REGION Network 9
   RUNG wire#powerrail
      Move(in := #AccumZnSpacing, out1 => #AccumSpacingEcho)
      Move(in := #ProductZoneSpacing, out1 => #ProdZoneSpacingEcho)
   END_RUNG
   // the same network as SCL:
   #AccumSpacingEcho := #AccumZnSpacing;
   #ProdZoneSpacingEcho := #ProductZoneSpacing;
END_REGION

REGION Network 10
   RUNG wire#powerrail
      { S7_Templates := "SrcType := Int" } NE_Contact(in1 := "EMS".Zone[#Zone].CarrierZnStatus[#MaxCarriers].CarrierNumber, in2 := 0)
      Coil( #ZoneFull )
   END_RUNG
   // the same network as SCL:
   #ZoneFull := "EMS".Zone[#Zone].CarrierZnStatus[#MaxCarriers].CarrierNumber <> 0;
END_REGION

REGION Network 11
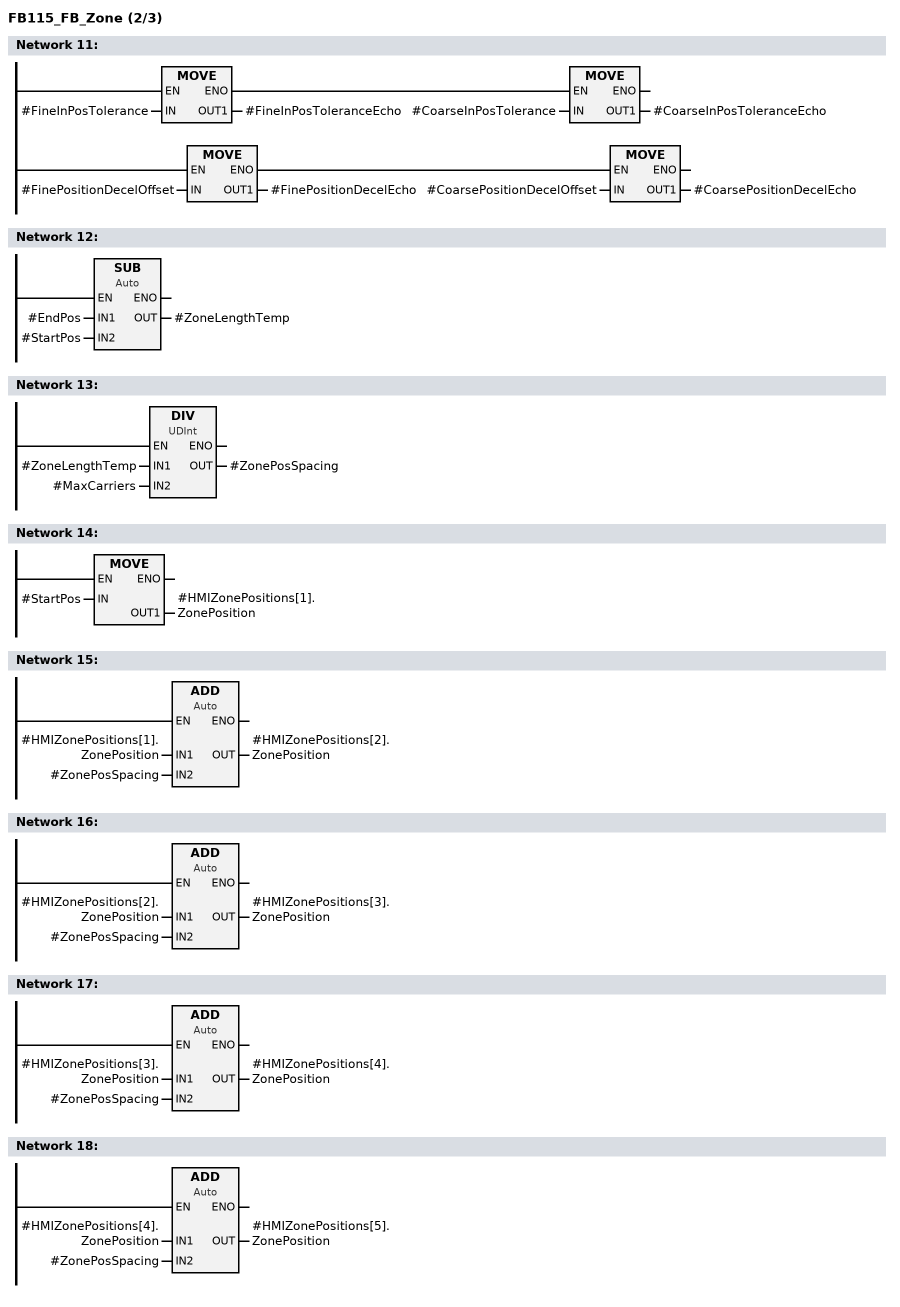
   RUNG wire#powerrail
      Move(in := #FineInPosTolerance, out1 => #FineInPosToleranceEcho)
      Move(in := #CoarseInPosTolerance, out1 => #CoarseInPosToleranceEcho)
   END_RUNG
   RUNG wire#powerrail
      Move(in := #FinePositionDecelOffset, out1 => #FinePositionDecelEcho)
      Move(in := #CoarsePositionDecelOffset, out1 => #CoarsePositionDecelEcho)
   END_RUNG
   // the same network as SCL:
   #FineInPosToleranceEcho := #FineInPosTolerance;
   #CoarseInPosToleranceEcho := #CoarseInPosTolerance;
   #FinePositionDecelEcho := #FinePositionDecelOffset;
   #CoarsePositionDecelEcho := #CoarsePositionDecelOffset;
END_REGION

REGION Network 12
   RUNG wire#powerrail
      Sub(in1 := #EndPos, in2 := #StartPos, out => #ZoneLengthTemp)
   END_RUNG
   // the same network as SCL:
   #ZoneLengthTemp := #EndPos - #StartPos;
END_REGION

REGION Network 13
   RUNG wire#powerrail
      { S7_Templates := "SrcType := UDInt" } Div(in1 := #ZoneLengthTemp, in2 := #MaxCarriers, out => #ZonePosSpacing)
   END_RUNG
   // the same network as SCL:
   #ZonePosSpacing := #ZoneLengthTemp / #MaxCarriers;
END_REGION

REGION Network 14
   RUNG wire#powerrail
      Move(in := #StartPos, out1 => #HMIZonePositions[1].ZonePosition)
   END_RUNG
   // the same network as SCL:
   #HMIZonePositions[1].ZonePosition := #StartPos;
END_REGION

REGION Network 15
   RUNG wire#powerrail
      Add(in1 := #HMIZonePositions[1].ZonePosition, in2 := #ZonePosSpacing, out => #HMIZonePositions[2].ZonePosition)
   END_RUNG
   // the same network as SCL:
   #HMIZonePositions[2].ZonePosition := #HMIZonePositions[1].ZonePosition + #ZonePosSpacing;
END_REGION

REGION Network 16
   RUNG wire#powerrail
      Add(in1 := #HMIZonePositions[2].ZonePosition, in2 := #ZonePosSpacing, out => #HMIZonePositions[3].ZonePosition)
   END_RUNG
   // the same network as SCL:
   #HMIZonePositions[3].ZonePosition := #HMIZonePositions[2].ZonePosition + #ZonePosSpacing;
END_REGION

REGION Network 17
   RUNG wire#powerrail
      Add(in1 := #HMIZonePositions[3].ZonePosition, in2 := #ZonePosSpacing, out => #HMIZonePositions[4].ZonePosition)
   END_RUNG
   // the same network as SCL:
   #HMIZonePositions[4].ZonePosition := #HMIZonePositions[3].ZonePosition + #ZonePosSpacing;
END_REGION

REGION Network 18
   RUNG wire#powerrail
      Add(in1 := #HMIZonePositions[4].ZonePosition, in2 := #ZonePosSpacing, out => #HMIZonePositions[5].ZonePosition)
   END_RUNG
   // the same network as SCL:
   #HMIZonePositions[5].ZonePosition := #HMIZonePositions[4].ZonePosition + #ZonePosSpacing;
END_REGION

REGION Network 19
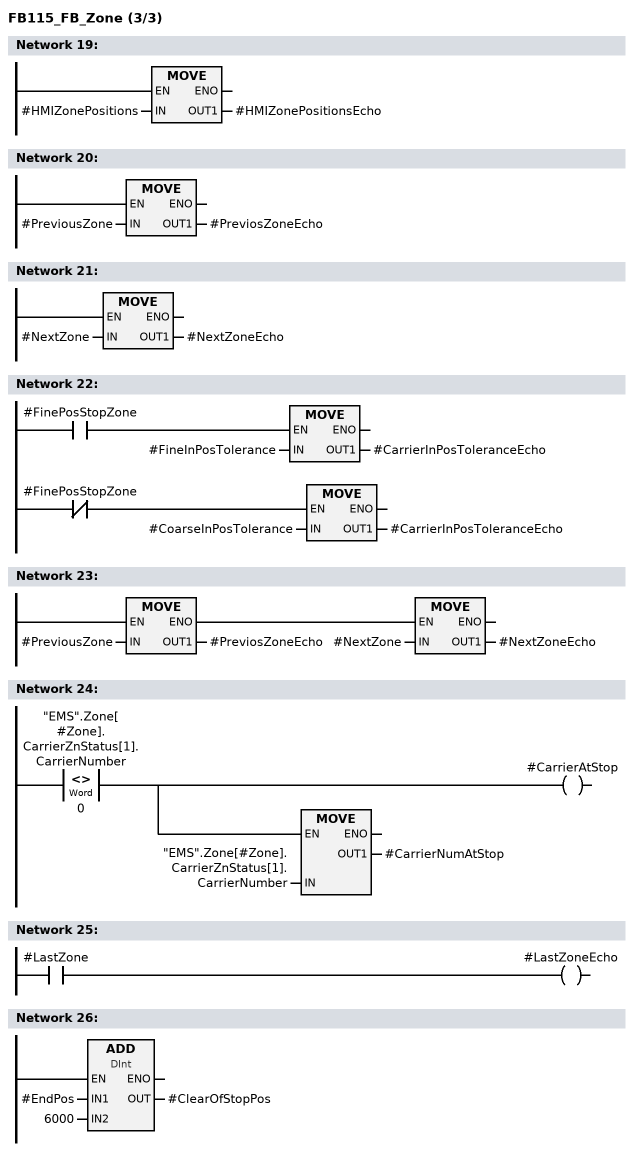
   RUNG wire#powerrail
      Move(in := #HMIZonePositions, out1 => #HMIZonePositionsEcho)
   END_RUNG
   // the same network as SCL:
   #HMIZonePositionsEcho := #HMIZonePositions;
END_REGION

REGION Network 20
   RUNG wire#powerrail
      Move(in := #PreviousZone, out1 => #PreviosZoneEcho)
   END_RUNG
   // the same network as SCL:
   #PreviosZoneEcho := #PreviousZone;
END_REGION

REGION Network 21
   RUNG wire#powerrail
      Move(in := #NextZone, out1 => #NextZoneEcho)
   END_RUNG
   // the same network as SCL:
   #NextZoneEcho := #NextZone;
END_REGION

REGION Network 22
   RUNG wire#powerrail
      Contact( #FinePosStopZone )
      Move(in := #FineInPosTolerance, out1 => #CarrierInPosToleranceEcho)
   END_RUNG
   RUNG wire#powerrail
      I_Contact( #FinePosStopZone )
      Move(in := #CoarseInPosTolerance, out1 => #CarrierInPosToleranceEcho)
   END_RUNG
   // the same network as SCL:
   IF #FinePosStopZone THEN #CarrierInPosToleranceEcho := #FineInPosTolerance; END_IF;
   IF NOT #FinePosStopZone THEN #CarrierInPosToleranceEcho := #CoarseInPosTolerance; END_IF;
END_REGION

REGION Network 23
   RUNG wire#powerrail
      Move(in := #PreviousZone, out1 => #PreviosZoneEcho)
      Move(in := #NextZone, out1 => #NextZoneEcho)
   END_RUNG
   // the same network as SCL:
   #PreviosZoneEcho := #PreviousZone;
   #NextZoneEcho := #NextZone;
END_REGION

REGION Network 24
   RUNG wire#powerrail
      { S7_Templates := "SrcType := Word" } NE_Contact(in1 := "EMS".Zone[#Zone].CarrierZnStatus[1].CarrierNumber, in2 := 0)
      wire#w1
      Coil( #CarrierAtStop )
   END_RUNG
   RUNG wire#w1
      Move(in := "EMS".Zone[#Zone].CarrierZnStatus[1].CarrierNumber, out1 => #CarrierNumAtStop)
   END_RUNG
   // the same network as SCL:
   #CarrierAtStop := "EMS".Zone[#Zone].CarrierZnStatus[1].CarrierNumber <> 0;
   IF #CarrierAtStop THEN #CarrierNumAtStop := "EMS".Zone[#Zone].CarrierZnStatus[1].CarrierNumber; END_IF;
END_REGION

REGION Network 25
   RUNG wire#powerrail
      Contact( #LastZone )
      Coil( #LastZoneEcho )
   END_RUNG
   // the same network as SCL:
   #LastZoneEcho := #LastZone;
END_REGION

REGION Network 26
   RUNG wire#powerrail
      { S7_Templates := "SrcType := DInt" } Add(in1 := #EndPos, in2 := 6000, out => #ClearOfStopPos)
   END_RUNG
   // the same network as SCL:
   #ClearOfStopPos := #EndPos + 6000;
END_REGION
END_FUNCTION_BLOCK

FUNCTION_BLOCK "FB116_FB_ZonePositionArrayTrafficCop"   // FB116, LAD
{ S7_Optimized_Access := 'FALSE' }
VERSION : 0.1
   VAR_INPUT
      Zone : Int := 1;
      CarrierZnArrayPos : Int;
   END_VAR
   VAR_OUTPUT
      MoveFwd : Bool;
      Speed : Word;
      TCZnPosnArray : "UDT_TrafficCopZoneStructure";
   END_VAR
   VAR
      CarNumZnPos : Array[0..99] of Int;
      TrafficCopCarrierZnBufferOut : Array[0..30] of "UDT_TrafficCop";
      "Zn-Pos2CarrierNumTemp" : Int;
      Zone1TrafficCopStructure : Struct
         CommandPosition : Word;
         InPositionTolerance : Word;
         CommandPositionUpperLimit : Word;
         CommandPositionLowerLimit : Word;
         AtCommandPos : Bool;
      END_STRUCT;
      SectionComment : Bool;
      NextCarrierZnArrayPos : Int;
   END_VAR
BEGIN

REGION Network 1: Section Comment-Section Logic for Current Carrier number in Position 1 thru Max Carrier in Zone Position Array
   // Section Logic for Current Carrier number in Position 1 - Max Carrier in Zone Position Array
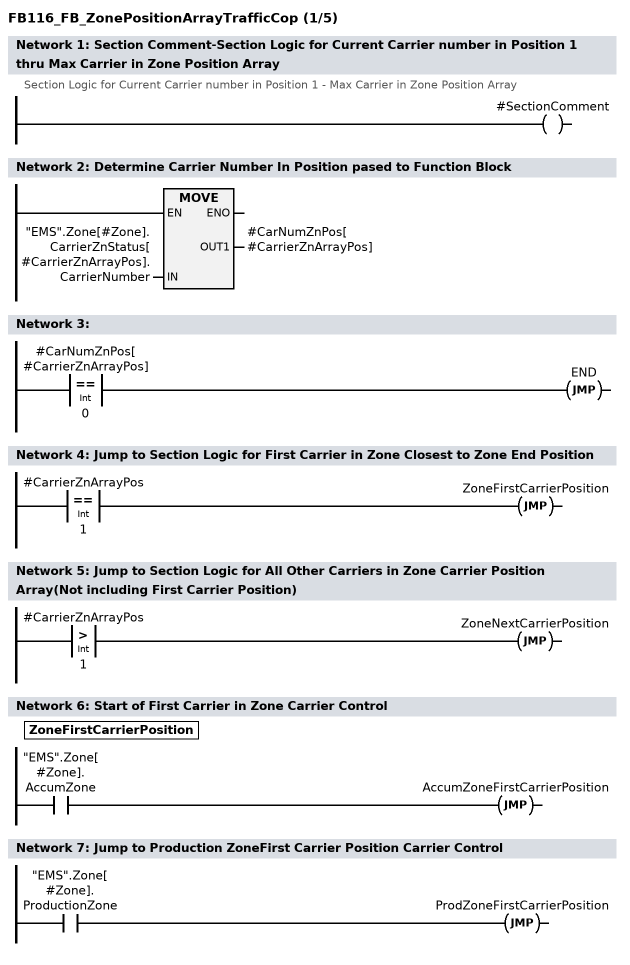
   RUNG wire#powerrail
      Coil( #SectionComment )
   END_RUNG
   // the same network as SCL:
   #SectionComment := TRUE;
END_REGION

REGION Network 2: Determine Carrier Number In Position pased to Function Block
   RUNG wire#powerrail
      Move(in := "EMS".Zone[#Zone].CarrierZnStatus[#CarrierZnArrayPos].CarrierNumber, out1 => #CarNumZnPos[#CarrierZnArrayPos])
   END_RUNG
   // the same network as SCL:
   #CarNumZnPos[#CarrierZnArrayPos] := "EMS".Zone[#Zone].CarrierZnStatus[#CarrierZnArrayPos].CarrierNumber;
END_REGION

REGION Network 3
   RUNG wire#powerrail
      { S7_Templates := "SrcType := Int" } EQ_Contact(in1 := #CarNumZnPos[#CarrierZnArrayPos], in2 := 0)
      JumpCoil( END )
   END_RUNG
   // the same network as SCL:
   IF #CarNumZnPos[#CarrierZnArrayPos] = 0 THEN GOTO END; END_IF;
END_REGION

REGION Network 4: Jump to Section Logic for First Carrier in Zone Closest to Zone End Position
   RUNG wire#powerrail
      { S7_Templates := "SrcType := Int" } EQ_Contact(in1 := #CarrierZnArrayPos, in2 := 1)
      JumpCoil( ZoneFirstCarrierPosition )
   END_RUNG
   // the same network as SCL:
   IF #CarrierZnArrayPos = 1 THEN GOTO ZoneFirstCarrierPosition; END_IF;
END_REGION

REGION Network 5: Jump to Section Logic for All Other Carriers in Zone Carrier Position Array(Not including First Carrier Position)
   RUNG wire#powerrail
      { S7_Templates := "SrcType := Int" } GT_Contact(in1 := #CarrierZnArrayPos, in2 := 1)
      JumpCoil( ZoneNextCarrierPosition )
   END_RUNG
   // the same network as SCL:
   IF #CarrierZnArrayPos > 1 THEN GOTO ZoneNextCarrierPosition; END_IF;
END_REGION

REGION Network 6: Start of First Carrier in Zone Carrier Control
   Label( ZoneFirstCarrierPosition )
   RUNG wire#powerrail
      Contact( "EMS".Zone[#Zone].AccumZone )
      JumpCoil( AccumZoneFirstCarrierPosition )
   END_RUNG
   // the same network as SCL:
   ZoneFirstCarrierPosition:
   IF "EMS".Zone[#Zone].AccumZone THEN GOTO AccumZoneFirstCarrierPosition; END_IF;
END_REGION

REGION Network 7: Jump to Production ZoneFirst Carrier Position Carrier Control
   RUNG wire#powerrail
      Contact( "EMS".Zone[#Zone].ProductionZone )
      JumpCoil( ProdZoneFirstCarrierPosition )
   END_RUNG
   // the same network as SCL:
   IF "EMS".Zone[#Zone].ProductionZone THEN GOTO ProdZoneFirstCarrierPosition; END_IF;
END_REGION

REGION Network 8: Position Carrier Control First Carrier in Accumulation Zone
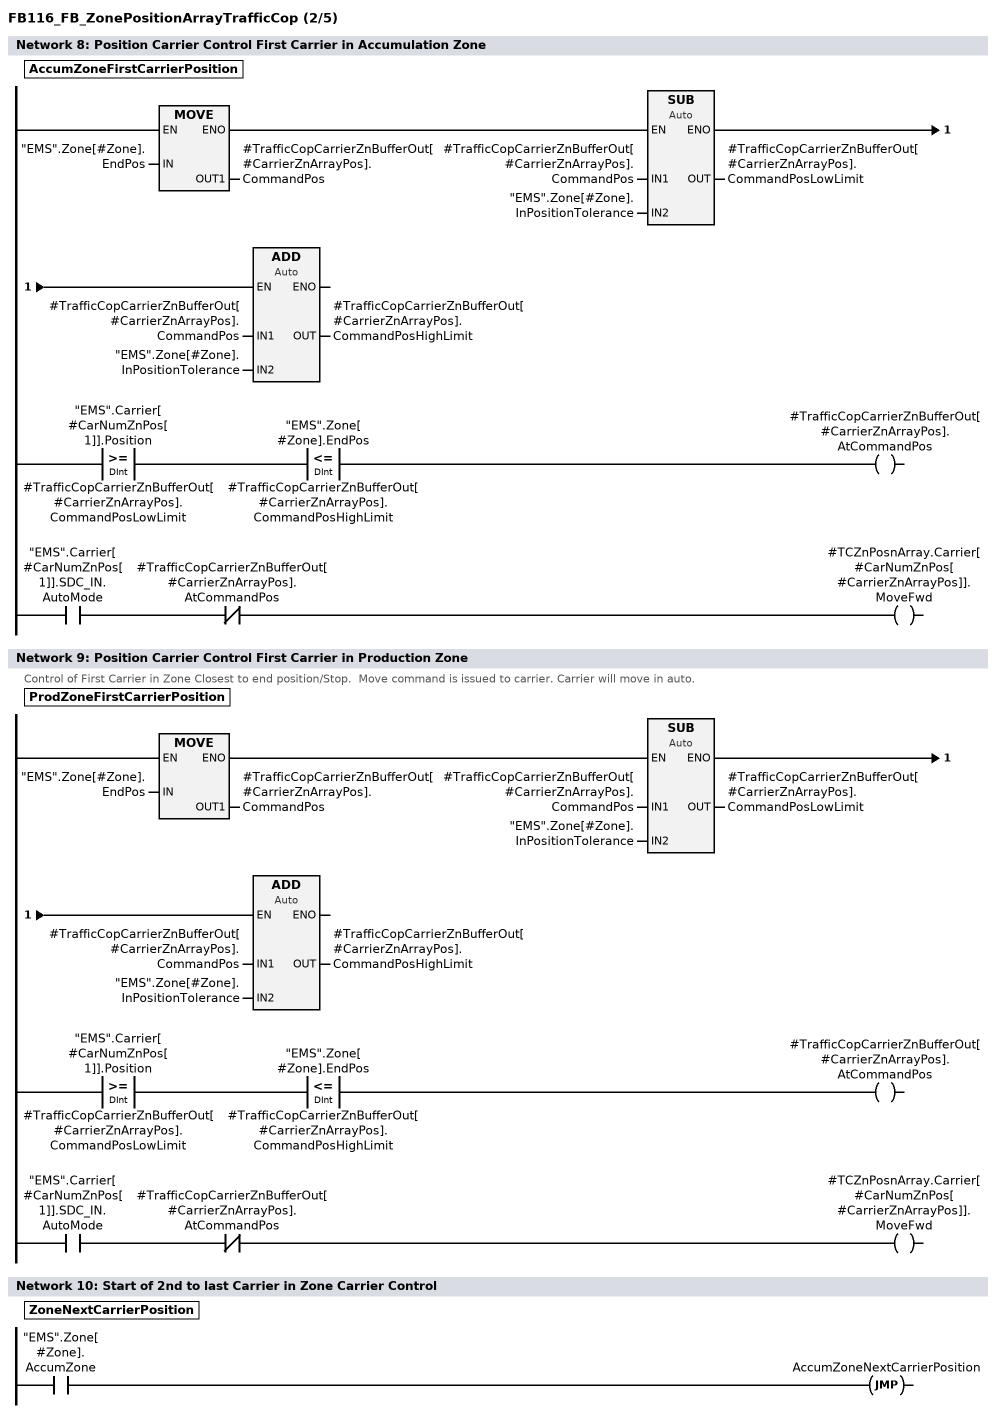
   Label( AccumZoneFirstCarrierPosition )
   RUNG wire#powerrail
      Move(in := "EMS".Zone[#Zone].EndPos, out1 => #TrafficCopCarrierZnBufferOut[#CarrierZnArrayPos].CommandPos)
      Sub(in1 := #TrafficCopCarrierZnBufferOut[#CarrierZnArrayPos].CommandPos, in2 := "EMS".Zone[#Zone].InPositionTolerance, out => #TrafficCopCarrierZnBufferOut[#CarrierZnArrayPos].CommandPosLowLimit)
      Add(in1 := #TrafficCopCarrierZnBufferOut[#CarrierZnArrayPos].CommandPos, in2 := "EMS".Zone[#Zone].InPositionTolerance, out => #TrafficCopCarrierZnBufferOut[#CarrierZnArrayPos].CommandPosHighLimit)
   END_RUNG
   RUNG wire#powerrail
      { S7_Templates := "SrcType := DInt" } GE_Contact(in1 := "EMS".Carrier[#CarNumZnPos[1]].Position, in2 := #TrafficCopCarrierZnBufferOut[#CarrierZnArrayPos].CommandPosLowLimit)
      { S7_Templates := "SrcType := DInt" } LE_Contact(in1 := "EMS".Zone[#Zone].EndPos, in2 := #TrafficCopCarrierZnBufferOut[#CarrierZnArrayPos].CommandPosHighLimit)
      Coil( #TrafficCopCarrierZnBufferOut[#CarrierZnArrayPos].AtCommandPos )
   END_RUNG
   RUNG wire#powerrail
      Contact( "EMS".Carrier[#CarNumZnPos[1]].SDC_IN.AutoMode )
      I_Contact( #TrafficCopCarrierZnBufferOut[#CarrierZnArrayPos].AtCommandPos )
      Coil( #TCZnPosnArray.Carrier[#CarNumZnPos[#CarrierZnArrayPos]].MoveFwd )
   END_RUNG
   // the same network as SCL:
   AccumZoneFirstCarrierPosition:
   #TrafficCopCarrierZnBufferOut[#CarrierZnArrayPos].CommandPos := "EMS".Zone[#Zone].EndPos;
   #TrafficCopCarrierZnBufferOut[#CarrierZnArrayPos].CommandPosLowLimit := #TrafficCopCarrierZnBufferOut[#CarrierZnArrayPos].CommandPos - "EMS".Zone[#Zone].InPositionTolerance;
   #TrafficCopCarrierZnBufferOut[#CarrierZnArrayPos].CommandPosHighLimit := #TrafficCopCarrierZnBufferOut[#CarrierZnArrayPos].CommandPos + "EMS".Zone[#Zone].InPositionTolerance;
   #TrafficCopCarrierZnBufferOut[#CarrierZnArrayPos].AtCommandPos := ("EMS".Carrier[#CarNumZnPos[1]].Position >= #TrafficCopCarrierZnBufferOut[#CarrierZnArrayPos].CommandPosLowLimit) AND ("EMS".Zone[#Zone].EndPos <= #TrafficCopCarrierZnBufferOut[#CarrierZnArrayPos].CommandPosHighLimit);
   #TCZnPosnArray.Carrier[#CarNumZnPos[#CarrierZnArrayPos]].MoveFwd := "EMS".Carrier[#CarNumZnPos[1]].SDC_IN.AutoMode AND NOT #TrafficCopCarrierZnBufferOut[#CarrierZnArrayPos].AtCommandPos;
END_REGION

REGION Network 9: Position Carrier Control First Carrier in Production Zone
   // Control of First Carrier in Zone Closest to end position/Stop.  Move command is issued to carrier. Carrier will move in auto.
   Label( ProdZoneFirstCarrierPosition )
   RUNG wire#powerrail
      Move(in := "EMS".Zone[#Zone].EndPos, out1 => #TrafficCopCarrierZnBufferOut[#CarrierZnArrayPos].CommandPos)
      Sub(in1 := #TrafficCopCarrierZnBufferOut[#CarrierZnArrayPos].CommandPos, in2 := "EMS".Zone[#Zone].InPositionTolerance, out => #TrafficCopCarrierZnBufferOut[#CarrierZnArrayPos].CommandPosLowLimit)
      Add(in1 := #TrafficCopCarrierZnBufferOut[#CarrierZnArrayPos].CommandPos, in2 := "EMS".Zone[#Zone].InPositionTolerance, out => #TrafficCopCarrierZnBufferOut[#CarrierZnArrayPos].CommandPosHighLimit)
   END_RUNG
   RUNG wire#powerrail
      { S7_Templates := "SrcType := DInt" } GE_Contact(in1 := "EMS".Carrier[#CarNumZnPos[1]].Position, in2 := #TrafficCopCarrierZnBufferOut[#CarrierZnArrayPos].CommandPosLowLimit)
      { S7_Templates := "SrcType := DInt" } LE_Contact(in1 := "EMS".Zone[#Zone].EndPos, in2 := #TrafficCopCarrierZnBufferOut[#CarrierZnArrayPos].CommandPosHighLimit)
      Coil( #TrafficCopCarrierZnBufferOut[#CarrierZnArrayPos].AtCommandPos )
   END_RUNG
   RUNG wire#powerrail
      Contact( "EMS".Carrier[#CarNumZnPos[1]].SDC_IN.AutoMode )
      I_Contact( #TrafficCopCarrierZnBufferOut[#CarrierZnArrayPos].AtCommandPos )
      Coil( #TCZnPosnArray.Carrier[#CarNumZnPos[#CarrierZnArrayPos]].MoveFwd )
   END_RUNG
   // the same network as SCL:
   ProdZoneFirstCarrierPosition:
   #TrafficCopCarrierZnBufferOut[#CarrierZnArrayPos].CommandPos := "EMS".Zone[#Zone].EndPos;
   #TrafficCopCarrierZnBufferOut[#CarrierZnArrayPos].CommandPosLowLimit := #TrafficCopCarrierZnBufferOut[#CarrierZnArrayPos].CommandPos - "EMS".Zone[#Zone].InPositionTolerance;
   #TrafficCopCarrierZnBufferOut[#CarrierZnArrayPos].CommandPosHighLimit := #TrafficCopCarrierZnBufferOut[#CarrierZnArrayPos].CommandPos + "EMS".Zone[#Zone].InPositionTolerance;
   #TrafficCopCarrierZnBufferOut[#CarrierZnArrayPos].AtCommandPos := ("EMS".Carrier[#CarNumZnPos[1]].Position >= #TrafficCopCarrierZnBufferOut[#CarrierZnArrayPos].CommandPosLowLimit) AND ("EMS".Zone[#Zone].EndPos <= #TrafficCopCarrierZnBufferOut[#CarrierZnArrayPos].CommandPosHighLimit);
   #TCZnPosnArray.Carrier[#CarNumZnPos[#CarrierZnArrayPos]].MoveFwd := "EMS".Carrier[#CarNumZnPos[1]].SDC_IN.AutoMode AND NOT #TrafficCopCarrierZnBufferOut[#CarrierZnArrayPos].AtCommandPos;
END_REGION

REGION Network 10: Start of 2nd to last Carrier in Zone Carrier Control
   Label( ZoneNextCarrierPosition )
   RUNG wire#powerrail
      Contact( "EMS".Zone[#Zone].AccumZone )
      JumpCoil( AccumZoneNextCarrierPosition )
   END_RUNG
   // the same network as SCL:
   ZoneNextCarrierPosition:
   IF "EMS".Zone[#Zone].AccumZone THEN GOTO AccumZoneNextCarrierPosition; END_IF;
END_REGION

REGION Network 11: Jump to Production Zone 2nd to Last Carrier Position Carrier Control
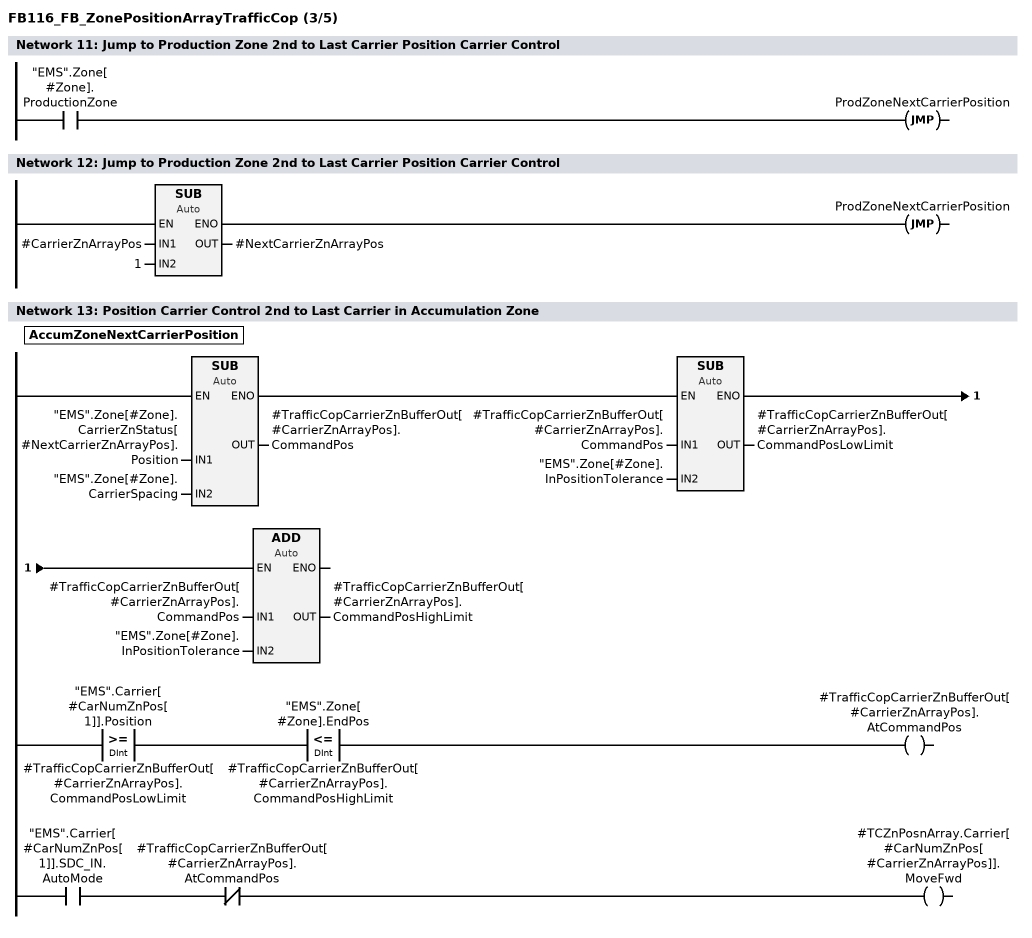
   RUNG wire#powerrail
      Contact( "EMS".Zone[#Zone].ProductionZone )
      JumpCoil( ProdZoneNextCarrierPosition )
   END_RUNG
   // the same network as SCL:
   IF "EMS".Zone[#Zone].ProductionZone THEN GOTO ProdZoneNextCarrierPosition; END_IF;
END_REGION

REGION Network 12: Jump to Production Zone 2nd to Last Carrier Position Carrier Control
   RUNG wire#powerrail
      Sub(in1 := #CarrierZnArrayPos, in2 := 1, out => #NextCarrierZnArrayPos)
      JumpCoil( ProdZoneNextCarrierPosition )
   END_RUNG
   // the same network as SCL:
   #NextCarrierZnArrayPos := #CarrierZnArrayPos - 1;
   GOTO ProdZoneNextCarrierPosition;
END_REGION

REGION Network 13: Position Carrier Control 2nd to Last Carrier in Accumulation Zone
   Label( AccumZoneNextCarrierPosition )
   RUNG wire#powerrail
      Sub(in1 := "EMS".Zone[#Zone].CarrierZnStatus[#NextCarrierZnArrayPos].Position, in2 := "EMS".Zone[#Zone].CarrierSpacing, out => #TrafficCopCarrierZnBufferOut[#CarrierZnArrayPos].CommandPos)
      Sub(in1 := #TrafficCopCarrierZnBufferOut[#CarrierZnArrayPos].CommandPos, in2 := "EMS".Zone[#Zone].InPositionTolerance, out => #TrafficCopCarrierZnBufferOut[#CarrierZnArrayPos].CommandPosLowLimit)
      Add(in1 := #TrafficCopCarrierZnBufferOut[#CarrierZnArrayPos].CommandPos, in2 := "EMS".Zone[#Zone].InPositionTolerance, out => #TrafficCopCarrierZnBufferOut[#CarrierZnArrayPos].CommandPosHighLimit)
   END_RUNG
   RUNG wire#powerrail
      { S7_Templates := "SrcType := DInt" } GE_Contact(in1 := "EMS".Carrier[#CarNumZnPos[1]].Position, in2 := #TrafficCopCarrierZnBufferOut[#CarrierZnArrayPos].CommandPosLowLimit)
      { S7_Templates := "SrcType := DInt" } LE_Contact(in1 := "EMS".Zone[#Zone].EndPos, in2 := #TrafficCopCarrierZnBufferOut[#CarrierZnArrayPos].CommandPosHighLimit)
      Coil( #TrafficCopCarrierZnBufferOut[#CarrierZnArrayPos].AtCommandPos )
   END_RUNG
   RUNG wire#powerrail
      Contact( "EMS".Carrier[#CarNumZnPos[1]].SDC_IN.AutoMode )
      I_Contact( #TrafficCopCarrierZnBufferOut[#CarrierZnArrayPos].AtCommandPos )
      Coil( #TCZnPosnArray.Carrier[#CarNumZnPos[#CarrierZnArrayPos]].MoveFwd )
   END_RUNG
   // the same network as SCL:
   AccumZoneNextCarrierPosition:
   #TrafficCopCarrierZnBufferOut[#CarrierZnArrayPos].CommandPos := "EMS".Zone[#Zone].CarrierZnStatus[#NextCarrierZnArrayPos].Position - "EMS".Zone[#Zone].CarrierSpacing;
   #TrafficCopCarrierZnBufferOut[#CarrierZnArrayPos].CommandPosLowLimit := #TrafficCopCarrierZnBufferOut[#CarrierZnArrayPos].CommandPos - "EMS".Zone[#Zone].InPositionTolerance;
   #TrafficCopCarrierZnBufferOut[#CarrierZnArrayPos].CommandPosHighLimit := #TrafficCopCarrierZnBufferOut[#CarrierZnArrayPos].CommandPos + "EMS".Zone[#Zone].InPositionTolerance;
   #TrafficCopCarrierZnBufferOut[#CarrierZnArrayPos].AtCommandPos := ("EMS".Carrier[#CarNumZnPos[1]].Position >= #TrafficCopCarrierZnBufferOut[#CarrierZnArrayPos].CommandPosLowLimit) AND ("EMS".Zone[#Zone].EndPos <= #TrafficCopCarrierZnBufferOut[#CarrierZnArrayPos].CommandPosHighLimit);
   #TCZnPosnArray.Carrier[#CarNumZnPos[#CarrierZnArrayPos]].MoveFwd := "EMS".Carrier[#CarNumZnPos[1]].SDC_IN.AutoMode AND NOT #TrafficCopCarrierZnBufferOut[#CarrierZnArrayPos].AtCommandPos;
END_REGION

REGION Network 14: Position Carrier Control 2nd to Last Carrier in Production Zone
   // Control of 2nd to Last Carrier in Zone Move to next zone with carrier spacing
   // .  Move command is issued to carrier. Carrier will move in auto.
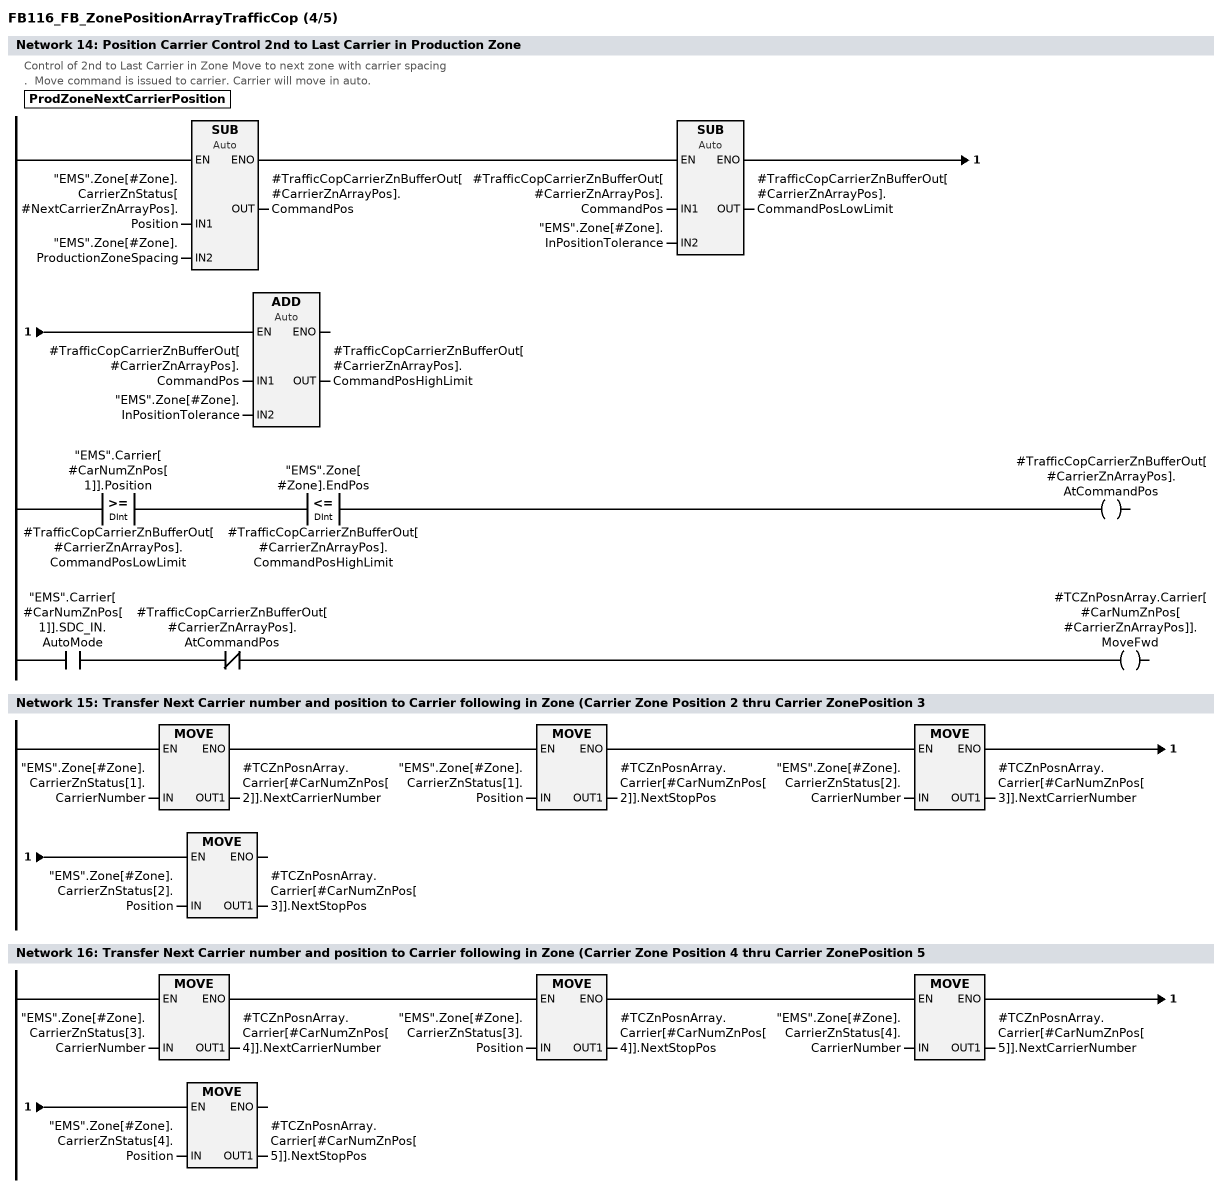
   Label( ProdZoneNextCarrierPosition )
   RUNG wire#powerrail
      Sub(in1 := "EMS".Zone[#Zone].CarrierZnStatus[#NextCarrierZnArrayPos].Position, in2 := "EMS".Zone[#Zone].ProductionZoneSpacing, out => #TrafficCopCarrierZnBufferOut[#CarrierZnArrayPos].CommandPos)
      Sub(in1 := #TrafficCopCarrierZnBufferOut[#CarrierZnArrayPos].CommandPos, in2 := "EMS".Zone[#Zone].InPositionTolerance, out => #TrafficCopCarrierZnBufferOut[#CarrierZnArrayPos].CommandPosLowLimit)
      Add(in1 := #TrafficCopCarrierZnBufferOut[#CarrierZnArrayPos].CommandPos, in2 := "EMS".Zone[#Zone].InPositionTolerance, out => #TrafficCopCarrierZnBufferOut[#CarrierZnArrayPos].CommandPosHighLimit)
   END_RUNG
   RUNG wire#powerrail
      { S7_Templates := "SrcType := DInt" } GE_Contact(in1 := "EMS".Carrier[#CarNumZnPos[1]].Position, in2 := #TrafficCopCarrierZnBufferOut[#CarrierZnArrayPos].CommandPosLowLimit)
      { S7_Templates := "SrcType := DInt" } LE_Contact(in1 := "EMS".Zone[#Zone].EndPos, in2 := #TrafficCopCarrierZnBufferOut[#CarrierZnArrayPos].CommandPosHighLimit)
      Coil( #TrafficCopCarrierZnBufferOut[#CarrierZnArrayPos].AtCommandPos )
   END_RUNG
   RUNG wire#powerrail
      Contact( "EMS".Carrier[#CarNumZnPos[1]].SDC_IN.AutoMode )
      I_Contact( #TrafficCopCarrierZnBufferOut[#CarrierZnArrayPos].AtCommandPos )
      Coil( #TCZnPosnArray.Carrier[#CarNumZnPos[#CarrierZnArrayPos]].MoveFwd )
   END_RUNG
   // the same network as SCL:
   ProdZoneNextCarrierPosition:
   #TrafficCopCarrierZnBufferOut[#CarrierZnArrayPos].CommandPos := "EMS".Zone[#Zone].CarrierZnStatus[#NextCarrierZnArrayPos].Position - "EMS".Zone[#Zone].ProductionZoneSpacing;
   #TrafficCopCarrierZnBufferOut[#CarrierZnArrayPos].CommandPosLowLimit := #TrafficCopCarrierZnBufferOut[#CarrierZnArrayPos].CommandPos - "EMS".Zone[#Zone].InPositionTolerance;
   #TrafficCopCarrierZnBufferOut[#CarrierZnArrayPos].CommandPosHighLimit := #TrafficCopCarrierZnBufferOut[#CarrierZnArrayPos].CommandPos + "EMS".Zone[#Zone].InPositionTolerance;
   #TrafficCopCarrierZnBufferOut[#CarrierZnArrayPos].AtCommandPos := ("EMS".Carrier[#CarNumZnPos[1]].Position >= #TrafficCopCarrierZnBufferOut[#CarrierZnArrayPos].CommandPosLowLimit) AND ("EMS".Zone[#Zone].EndPos <= #TrafficCopCarrierZnBufferOut[#CarrierZnArrayPos].CommandPosHighLimit);
   #TCZnPosnArray.Carrier[#CarNumZnPos[#CarrierZnArrayPos]].MoveFwd := "EMS".Carrier[#CarNumZnPos[1]].SDC_IN.AutoMode AND NOT #TrafficCopCarrierZnBufferOut[#CarrierZnArrayPos].AtCommandPos;
END_REGION

REGION Network 15: Transfer Next Carrier number and position to Carrier following in Zone (Carrier Zone Position 2 thru Carrier ZonePosition 3
   RUNG wire#powerrail
      Move(in := "EMS".Zone[#Zone].CarrierZnStatus[1].CarrierNumber, out1 => #TCZnPosnArray.Carrier[#CarNumZnPos[2]].NextCarrierNumber)
      Move(in := "EMS".Zone[#Zone].CarrierZnStatus[1].Position, out1 => #TCZnPosnArray.Carrier[#CarNumZnPos[2]].NextStopPos)
      Move(in := "EMS".Zone[#Zone].CarrierZnStatus[2].CarrierNumber, out1 => #TCZnPosnArray.Carrier[#CarNumZnPos[3]].NextCarrierNumber)
      Move(in := "EMS".Zone[#Zone].CarrierZnStatus[2].Position, out1 => #TCZnPosnArray.Carrier[#CarNumZnPos[3]].NextStopPos)
   END_RUNG
   // the same network as SCL:
   #TCZnPosnArray.Carrier[#CarNumZnPos[2]].NextCarrierNumber := "EMS".Zone[#Zone].CarrierZnStatus[1].CarrierNumber;
   #TCZnPosnArray.Carrier[#CarNumZnPos[2]].NextStopPos := "EMS".Zone[#Zone].CarrierZnStatus[1].Position;
   #TCZnPosnArray.Carrier[#CarNumZnPos[3]].NextCarrierNumber := "EMS".Zone[#Zone].CarrierZnStatus[2].CarrierNumber;
   #TCZnPosnArray.Carrier[#CarNumZnPos[3]].NextStopPos := "EMS".Zone[#Zone].CarrierZnStatus[2].Position;
END_REGION

REGION Network 16: Transfer Next Carrier number and position to Carrier following in Zone (Carrier Zone Position 4 thru Carrier ZonePosition 5
   RUNG wire#powerrail
      Move(in := "EMS".Zone[#Zone].CarrierZnStatus[3].CarrierNumber, out1 => #TCZnPosnArray.Carrier[#CarNumZnPos[4]].NextCarrierNumber)
      Move(in := "EMS".Zone[#Zone].CarrierZnStatus[3].Position, out1 => #TCZnPosnArray.Carrier[#CarNumZnPos[4]].NextStopPos)
      Move(in := "EMS".Zone[#Zone].CarrierZnStatus[4].CarrierNumber, out1 => #TCZnPosnArray.Carrier[#CarNumZnPos[5]].NextCarrierNumber)
      Move(in := "EMS".Zone[#Zone].CarrierZnStatus[4].Position, out1 => #TCZnPosnArray.Carrier[#CarNumZnPos[5]].NextStopPos)
   END_RUNG
   // the same network as SCL:
   #TCZnPosnArray.Carrier[#CarNumZnPos[4]].NextCarrierNumber := "EMS".Zone[#Zone].CarrierZnStatus[3].CarrierNumber;
   #TCZnPosnArray.Carrier[#CarNumZnPos[4]].NextStopPos := "EMS".Zone[#Zone].CarrierZnStatus[3].Position;
   #TCZnPosnArray.Carrier[#CarNumZnPos[5]].NextCarrierNumber := "EMS".Zone[#Zone].CarrierZnStatus[4].CarrierNumber;
   #TCZnPosnArray.Carrier[#CarNumZnPos[5]].NextStopPos := "EMS".Zone[#Zone].CarrierZnStatus[4].Position;
END_REGION

REGION Network 17: Transfer Next Carrier number and position to Carrier following in Zone (Carrier Zone Position 6 thru Carrier ZonePosition 7
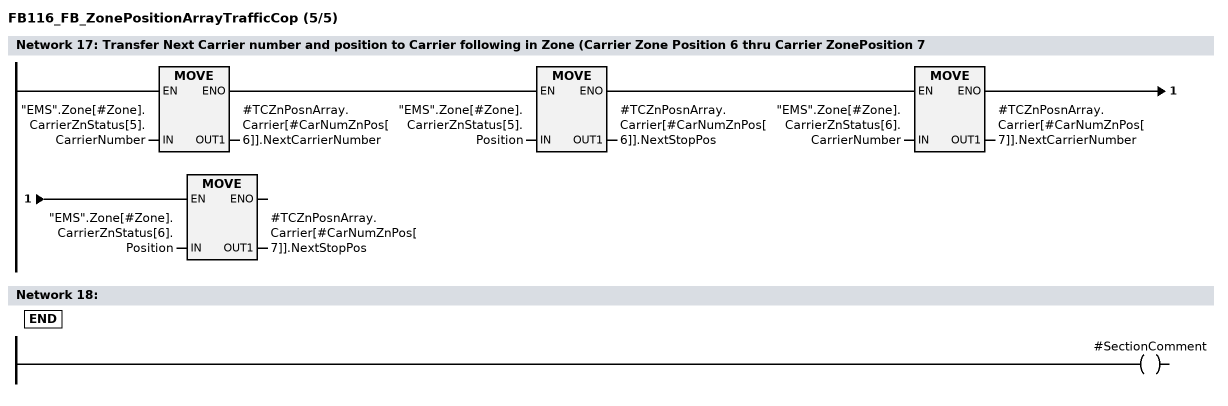
   RUNG wire#powerrail
      Move(in := "EMS".Zone[#Zone].CarrierZnStatus[5].CarrierNumber, out1 => #TCZnPosnArray.Carrier[#CarNumZnPos[6]].NextCarrierNumber)
      Move(in := "EMS".Zone[#Zone].CarrierZnStatus[5].Position, out1 => #TCZnPosnArray.Carrier[#CarNumZnPos[6]].NextStopPos)
      Move(in := "EMS".Zone[#Zone].CarrierZnStatus[6].CarrierNumber, out1 => #TCZnPosnArray.Carrier[#CarNumZnPos[7]].NextCarrierNumber)
      Move(in := "EMS".Zone[#Zone].CarrierZnStatus[6].Position, out1 => #TCZnPosnArray.Carrier[#CarNumZnPos[7]].NextStopPos)
   END_RUNG
   // the same network as SCL:
   #TCZnPosnArray.Carrier[#CarNumZnPos[6]].NextCarrierNumber := "EMS".Zone[#Zone].CarrierZnStatus[5].CarrierNumber;
   #TCZnPosnArray.Carrier[#CarNumZnPos[6]].NextStopPos := "EMS".Zone[#Zone].CarrierZnStatus[5].Position;
   #TCZnPosnArray.Carrier[#CarNumZnPos[7]].NextCarrierNumber := "EMS".Zone[#Zone].CarrierZnStatus[6].CarrierNumber;
   #TCZnPosnArray.Carrier[#CarNumZnPos[7]].NextStopPos := "EMS".Zone[#Zone].CarrierZnStatus[6].Position;
END_REGION

REGION Network 18
   Label( END )
   RUNG wire#powerrail
      Coil( #SectionComment )
   END_RUNG
   // the same network as SCL:
   END:
   #SectionComment := TRUE;
END_REGION
END_FUNCTION_BLOCK

FUNCTION_BLOCK "FB117_MapSDCOut_Carrier"   // FB117, LAD
{ S7_Optimized_Access := 'TRUE' }
VERSION : 0.1
   VAR_INPUT
      ZoneArray : Array[0..60] of "UDT_TC_SDCOutZone";
      Carrier : Int;
      Zone : Int;
   END_VAR
   VAR_OUTPUT
      DriveFwdCMD : Bool;
      AtCmdPos : Bool;
      NextStopPos : DWord;
      DriveCmdSpeed : Int;
      Zone_Echo : Int;
      Pos_Echo : DWord;
   END_VAR
   VAR
      CarrierArray : Array[0..99] of "UDT_TC_SDCOutCarrier";
   END_VAR
   VAR_TEMP   // added for the SCL form of the ladder/FBD networks
      _w1 : Bool;
   END_VAR
BEGIN

REGION Network 1
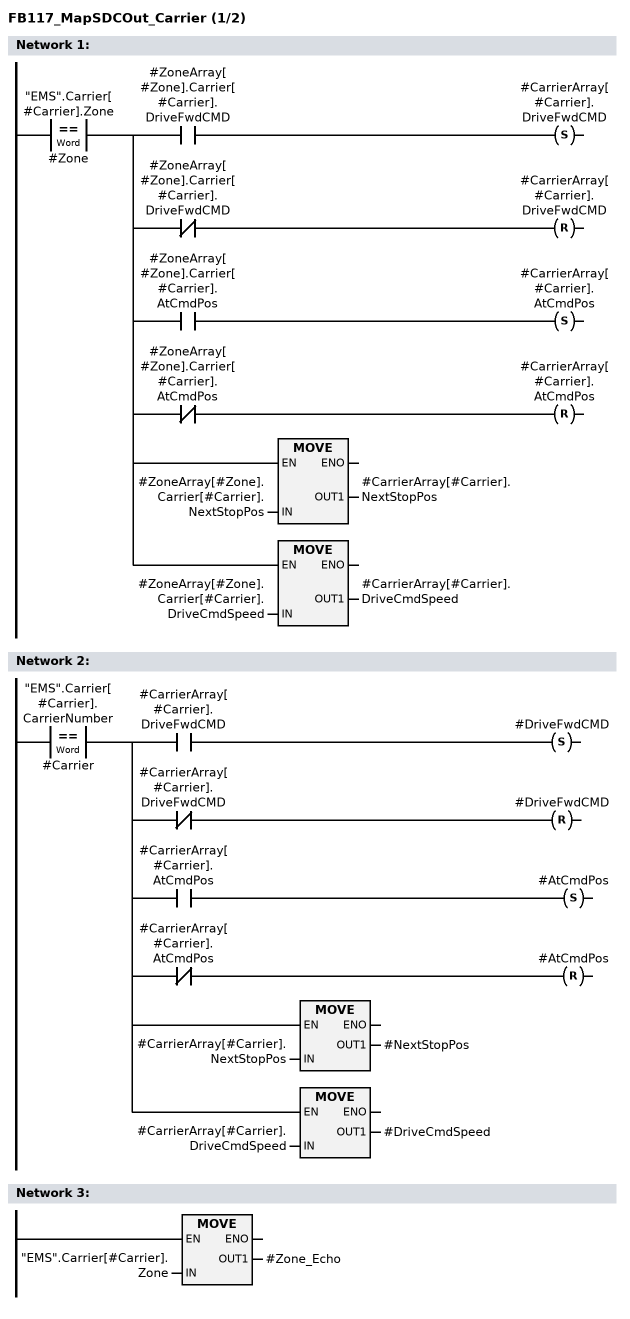
   RUNG wire#powerrail
      { S7_Templates := "SrcType := Word" } EQ_Contact(in1 := "EMS".Carrier[#Carrier].Zone, in2 := #Zone)
      wire#w1
      Contact( #ZoneArray[#Zone].Carrier[#Carrier].DriveFwdCMD )
      S_Coil( #CarrierArray[#Carrier].DriveFwdCMD )
   END_RUNG
   RUNG wire#w1
      I_Contact( #ZoneArray[#Zone].Carrier[#Carrier].DriveFwdCMD )
      R_Coil( #CarrierArray[#Carrier].DriveFwdCMD )
   END_RUNG
   RUNG wire#w1
      Contact( #ZoneArray[#Zone].Carrier[#Carrier].AtCmdPos )
      S_Coil( #CarrierArray[#Carrier].AtCmdPos )
   END_RUNG
   RUNG wire#w1
      I_Contact( #ZoneArray[#Zone].Carrier[#Carrier].AtCmdPos )
      R_Coil( #CarrierArray[#Carrier].AtCmdPos )
   END_RUNG
   RUNG wire#w1
      Move(in := #ZoneArray[#Zone].Carrier[#Carrier].NextStopPos, out1 => #CarrierArray[#Carrier].NextStopPos)
   END_RUNG
   RUNG wire#w1
      Move(in := #ZoneArray[#Zone].Carrier[#Carrier].DriveCmdSpeed, out1 => #CarrierArray[#Carrier].DriveCmdSpeed)
   END_RUNG
   // the same network as SCL:
   #_w1 := "EMS".Carrier[#Carrier].Zone = #Zone;
   IF #_w1 AND #ZoneArray[#Zone].Carrier[#Carrier].DriveFwdCMD THEN
       #CarrierArray[#Carrier].DriveFwdCMD := TRUE;
   END_IF;
   IF #_w1 AND NOT #ZoneArray[#Zone].Carrier[#Carrier].DriveFwdCMD THEN
       #CarrierArray[#Carrier].DriveFwdCMD := FALSE;
   END_IF;
   IF #_w1 AND #ZoneArray[#Zone].Carrier[#Carrier].AtCmdPos THEN
       #CarrierArray[#Carrier].AtCmdPos := TRUE;
   END_IF;
   IF #_w1 AND NOT #ZoneArray[#Zone].Carrier[#Carrier].AtCmdPos THEN
       #CarrierArray[#Carrier].AtCmdPos := FALSE;
   END_IF;
   IF #_w1 THEN
       #CarrierArray[#Carrier].NextStopPos := #ZoneArray[#Zone].Carrier[#Carrier].NextStopPos;
       #CarrierArray[#Carrier].DriveCmdSpeed := #ZoneArray[#Zone].Carrier[#Carrier].DriveCmdSpeed;
   END_IF;
END_REGION

REGION Network 2
   RUNG wire#powerrail
      { S7_Templates := "SrcType := Word" } EQ_Contact(in1 := "EMS".Carrier[#Carrier].CarrierNumber, in2 := #Carrier)
      wire#w1
      Contact( #CarrierArray[#Carrier].DriveFwdCMD )
      S_Coil( #DriveFwdCMD )
   END_RUNG
   RUNG wire#w1
      I_Contact( #CarrierArray[#Carrier].DriveFwdCMD )
      R_Coil( #DriveFwdCMD )
   END_RUNG
   RUNG wire#w1
      Contact( #CarrierArray[#Carrier].AtCmdPos )
      S_Coil( #AtCmdPos )
   END_RUNG
   RUNG wire#w1
      I_Contact( #CarrierArray[#Carrier].AtCmdPos )
      R_Coil( #AtCmdPos )
   END_RUNG
   RUNG wire#w1
      Move(in := #CarrierArray[#Carrier].NextStopPos, out1 => #NextStopPos)
   END_RUNG
   RUNG wire#w1
      Move(in := #CarrierArray[#Carrier].DriveCmdSpeed, out1 => #DriveCmdSpeed)
   END_RUNG
   // the same network as SCL:
   #_w1 := "EMS".Carrier[#Carrier].CarrierNumber = #Carrier;
   IF #_w1 AND #CarrierArray[#Carrier].DriveFwdCMD THEN #DriveFwdCMD := TRUE; END_IF;
   IF #_w1 AND NOT #CarrierArray[#Carrier].DriveFwdCMD THEN #DriveFwdCMD := FALSE; END_IF;
   IF #_w1 AND #CarrierArray[#Carrier].AtCmdPos THEN #AtCmdPos := TRUE; END_IF;
   IF #_w1 AND NOT #CarrierArray[#Carrier].AtCmdPos THEN #AtCmdPos := FALSE; END_IF;
   IF #_w1 THEN
       #NextStopPos := #CarrierArray[#Carrier].NextStopPos;
       #DriveCmdSpeed := #CarrierArray[#Carrier].DriveCmdSpeed;
   END_IF;
END_REGION
